ORGANIZATION_BLOCK "Cycle Execution"   // OB1, LAD
{ S7_Optimized_Access := 'FALSE' }
VERSION : 0.1
   VAR_TEMP
      TEMP0 : Byte;
      TEMP1 : Byte;
      TEMP2 : Byte;
      TEMP3 : Byte;
      TEMP4 : Byte;
      TEMP5 : Byte;
      TEMP6 : Int;
      TEMP7 : Int;
      TEMP8 : Int;
      TEMP9 : Date_And_Time;
      TEMP10 : DInt;
      TEMP11 : Int;
   END_VAR
   VAR_TEMP   // added for the SCL form of the ladder/FBD networks
      _w1 : Bool;
   END_VAR
BEGIN

REGION Network 1: -ALARMA
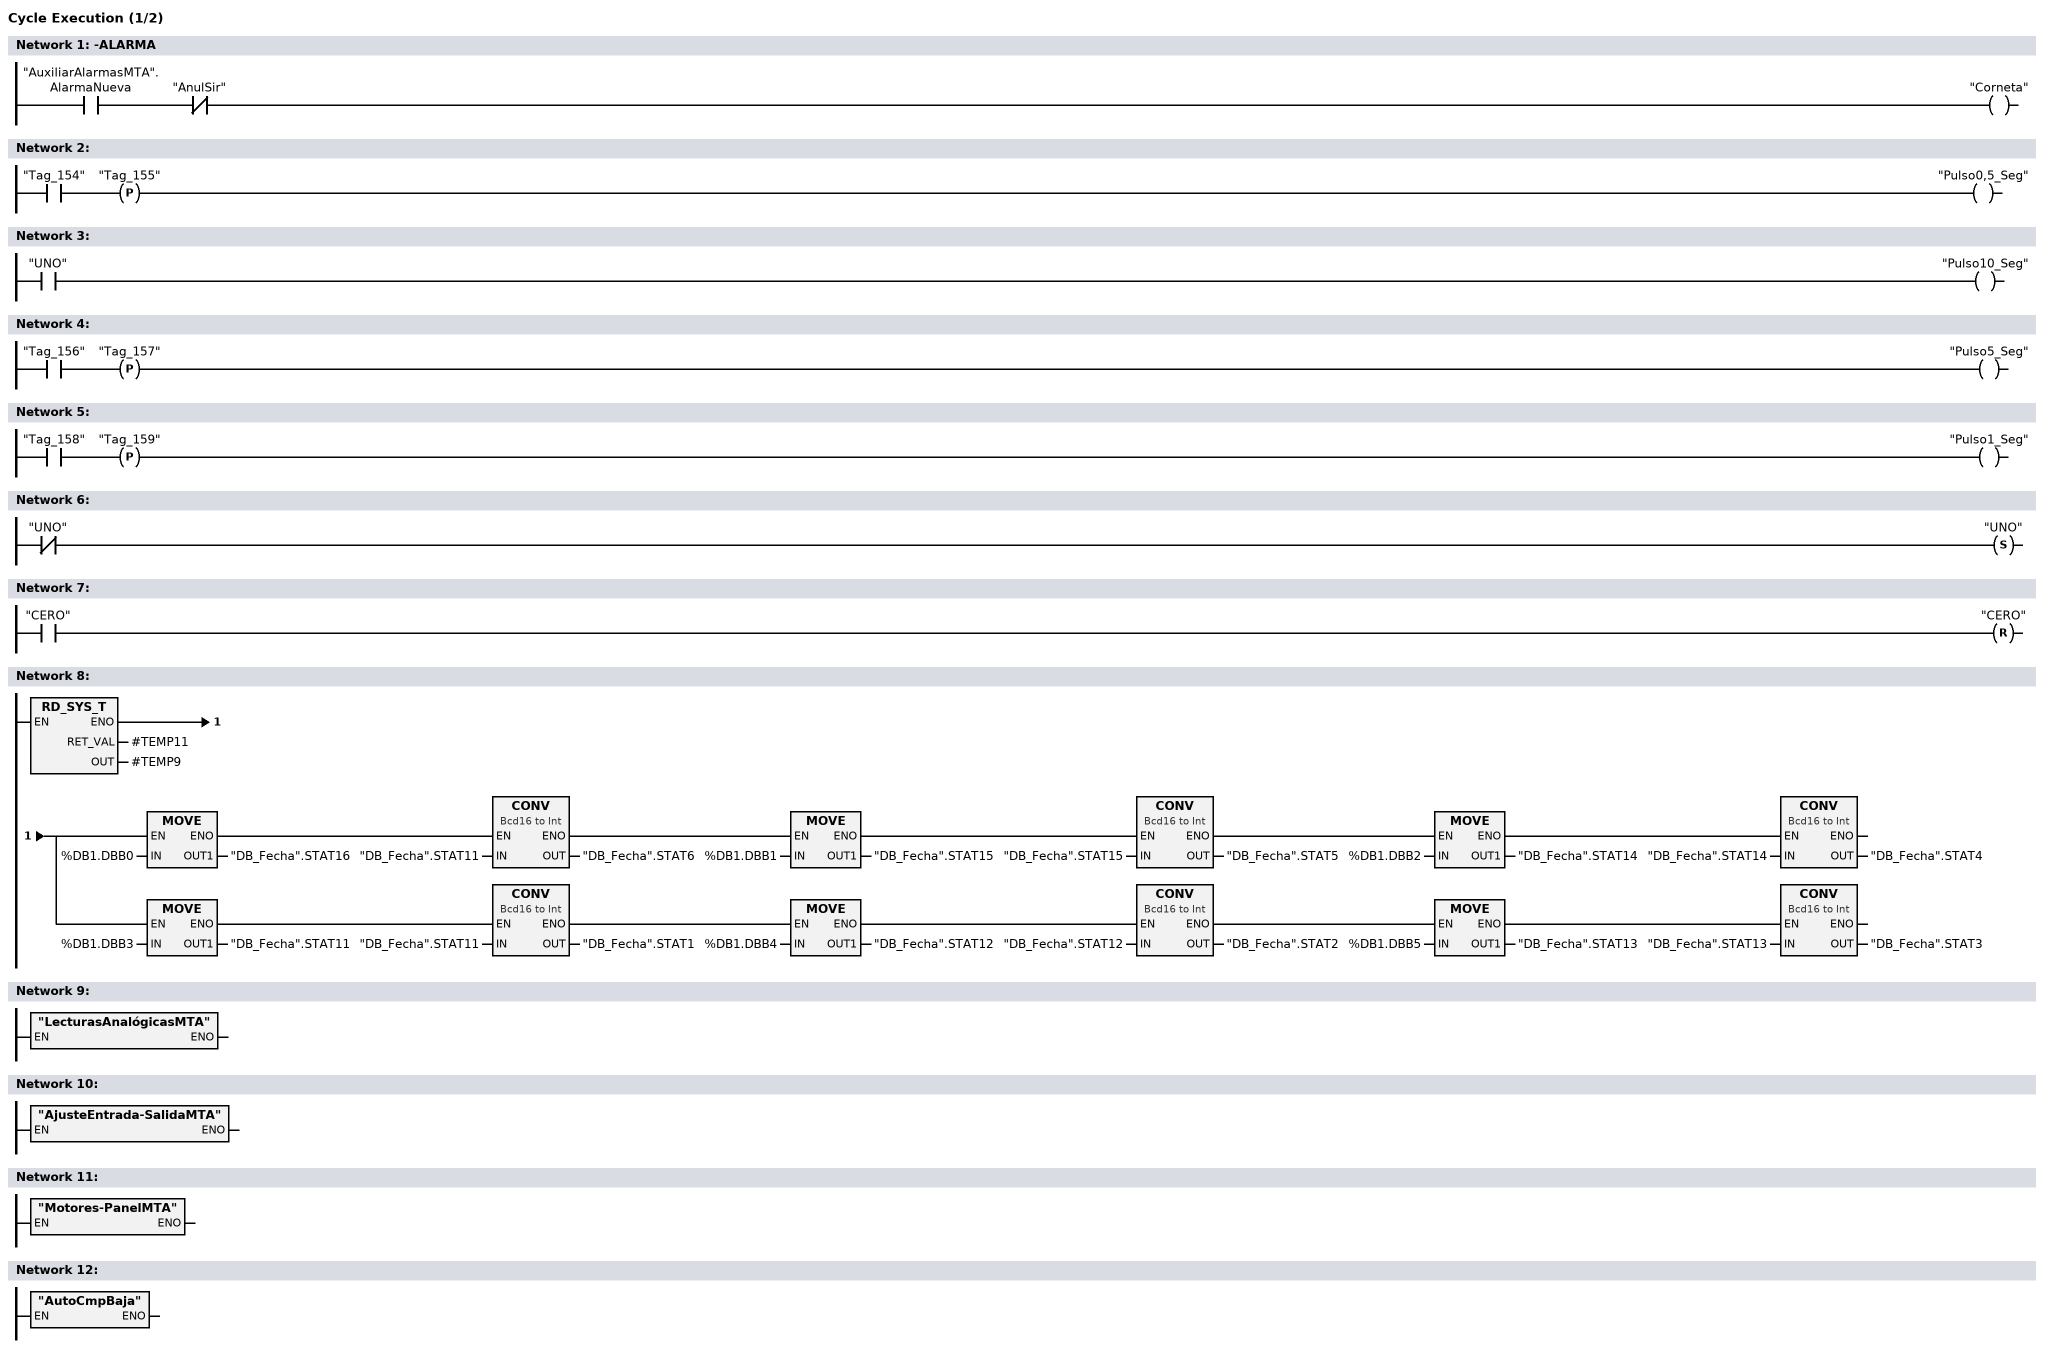
   RUNG wire#powerrail
      Contact( "AuxiliarAlarmasMTA".AlarmaNueva )
      I_Contact( "AnulSir" )
      Coil( "Corneta" )
   END_RUNG
   // the same network as SCL:
   "Corneta" := "AuxiliarAlarmasMTA".AlarmaNueva AND NOT "AnulSir";
END_REGION

REGION Network 2
   RUNG wire#powerrail
      Contact( "Tag_154" )
      P_Trig( "Tag_155" )
      Coil( "Pulso0,5_Seg" )
   END_RUNG
   // the same network as SCL:
   #_w1 := "Tag_154" AND NOT "Tag_155";   // rising edge
   "Tag_155" := "Tag_154";
   "Pulso0,5_Seg" := #_w1;
END_REGION

REGION Network 3
   RUNG wire#powerrail
      Contact( "UNO" )
      Coil( "Pulso10_Seg" )
   END_RUNG
   // the same network as SCL:
   "Pulso10_Seg" := "UNO";
END_REGION

REGION Network 4
   RUNG wire#powerrail
      Contact( "Tag_156" )
      P_Trig( "Tag_157" )
      Coil( "Pulso5_Seg" )
   END_RUNG
   // the same network as SCL:
   #_w1 := "Tag_156" AND NOT "Tag_157";   // rising edge
   "Tag_157" := "Tag_156";
   "Pulso5_Seg" := #_w1;
END_REGION

REGION Network 5
   RUNG wire#powerrail
      Contact( "Tag_158" )
      P_Trig( "Tag_159" )
      Coil( "Pulso1_Seg" )
   END_RUNG
   // the same network as SCL:
   #_w1 := "Tag_158" AND NOT "Tag_159";   // rising edge
   "Tag_159" := "Tag_158";
   "Pulso1_Seg" := #_w1;
END_REGION

REGION Network 6
   RUNG wire#powerrail
      I_Contact( "UNO" )
      S_Coil( "UNO" )
   END_RUNG
   // the same network as SCL:
   IF NOT "UNO" THEN "UNO" := TRUE; END_IF;
END_REGION

REGION Network 7
   RUNG wire#powerrail
      Contact( "CERO" )
      R_Coil( "CERO" )
   END_RUNG
   // the same network as SCL:
   IF "CERO" THEN "CERO" := FALSE; END_IF;
END_REGION

REGION Network 8
   // ENO of a box is taken as its EN; it also drops when the box reports an error
   #TEMP11 := RD_SYS_T(OUT => #TEMP9);
   "DB_Fecha".STAT16 := %DB1.DBB0;
   "DB_Fecha".STAT6 := BCD16_TO_INT("DB_Fecha".STAT11);
   "DB_Fecha".STAT15 := %DB1.DBB1;
   "DB_Fecha".STAT5 := BCD16_TO_INT("DB_Fecha".STAT15);
   "DB_Fecha".STAT14 := %DB1.DBB2;
   "DB_Fecha".STAT4 := BCD16_TO_INT("DB_Fecha".STAT14);
   "DB_Fecha".STAT11 := %DB1.DBB3;
   "DB_Fecha".STAT1 := BCD16_TO_INT("DB_Fecha".STAT11);
   "DB_Fecha".STAT12 := %DB1.DBB4;
   "DB_Fecha".STAT2 := BCD16_TO_INT("DB_Fecha".STAT12);
   "DB_Fecha".STAT13 := %DB1.DBB5;
   "DB_Fecha".STAT3 := BCD16_TO_INT("DB_Fecha".STAT13);
END_REGION

REGION Network 9
   RUNG wire#powerrail
      "LecturasAnalógicasMTA"()
   END_RUNG
   // the same network as SCL:
   "LecturasAnalógicasMTA"();
END_REGION

REGION Network 10
   RUNG wire#powerrail
      "AjusteEntrada-SalidaMTA"()
   END_RUNG
   // the same network as SCL:
   "AjusteEntrada-SalidaMTA"();
END_REGION

REGION Network 11
   RUNG wire#powerrail
      "Motores-PanelMTA"()
   END_RUNG
   // the same network as SCL:
   "Motores-PanelMTA"();
END_REGION

REGION Network 12
   RUNG wire#powerrail
      "AutoCmpBaja"()
   END_RUNG
   // the same network as SCL:
   "AutoCmpBaja"();
END_REGION

REGION Network 13
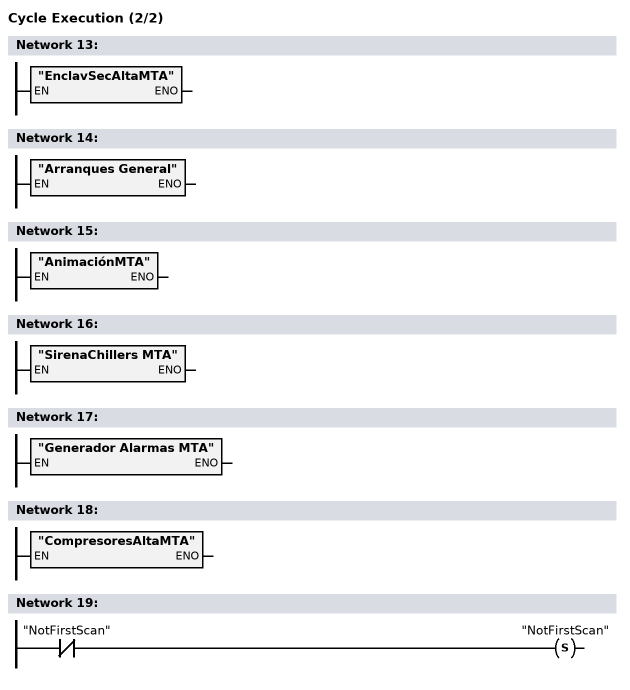
   RUNG wire#powerrail
      "EnclavSecAltaMTA"()
   END_RUNG
   // the same network as SCL:
   "EnclavSecAltaMTA"();
END_REGION

REGION Network 14
   RUNG wire#powerrail
      "Arranques General"()
   END_RUNG
   // the same network as SCL:
   "Arranques General"();
END_REGION

REGION Network 15
   RUNG wire#powerrail
      "AnimaciónMTA"()
   END_RUNG
   // the same network as SCL:
   "AnimaciónMTA"();
END_REGION

REGION Network 16
   RUNG wire#powerrail
      "SirenaChillers MTA"()
   END_RUNG
   // the same network as SCL:
   "SirenaChillers MTA"();
END_REGION

REGION Network 17
   RUNG wire#powerrail
      "Generador Alarmas MTA"()
   END_RUNG
   // the same network as SCL:
   "Generador Alarmas MTA"();
END_REGION

REGION Network 18
   RUNG wire#powerrail
      "CompresoresAltaMTA"()
   END_RUNG
   // the same network as SCL:
   "CompresoresAltaMTA"();
END_REGION

REGION Network 19
   RUNG wire#powerrail
      I_Contact( "NotFirstScan" )
      S_Coil( "NotFirstScan" )
   END_RUNG
   // the same network as SCL:
   IF NOT "NotFirstScan" THEN "NotFirstScan" := TRUE; END_IF;
END_REGION
END_ORGANIZATION_BLOCK

// folder: Alarmas

FUNCTION "SirenaChillers MTA" : Void   // FC7, LAD
{ S7_Optimized_Access := 'FALSE' }
VERSION : 0.1
BEGIN

REGION Network 1
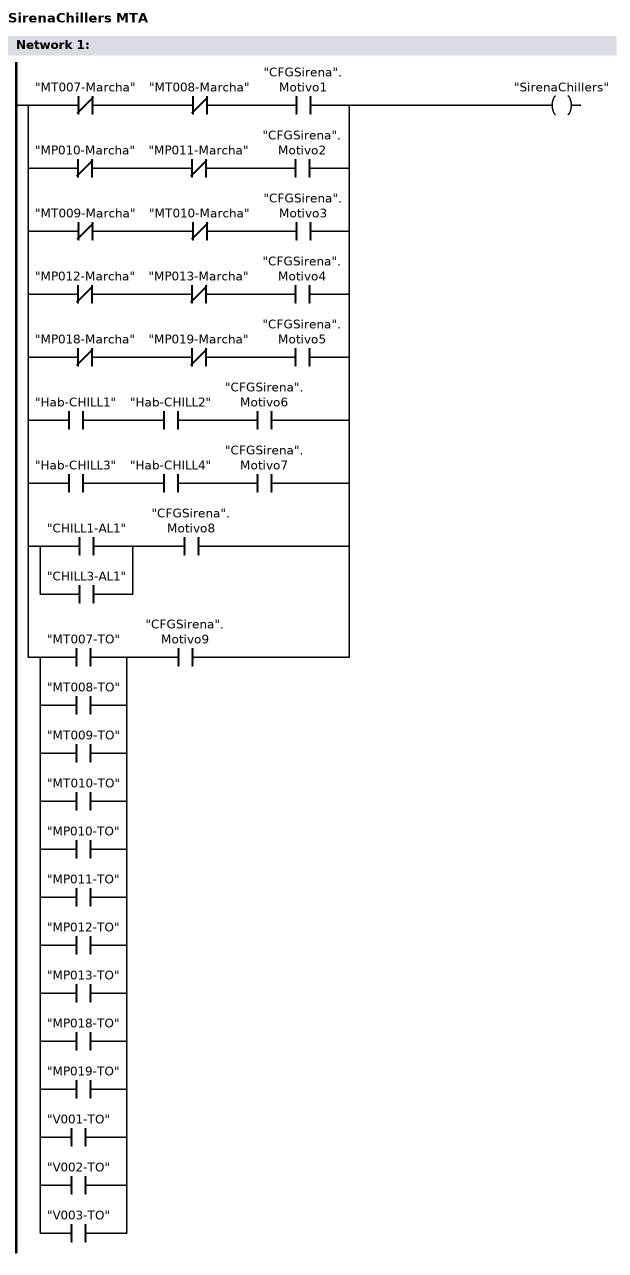
   RUNG wire#powerrail
      I_Contact( "MT007-Marcha" )
      I_Contact( "MT008-Marcha" )
      Contact( "CFGSirena".Motivo1 )
      wire#w1
      Coil( "SirenaChillers" )
   END_RUNG
   RUNG wire#powerrail
      I_Contact( "MP010-Marcha" )
      I_Contact( "MP011-Marcha" )
      Contact( "CFGSirena".Motivo2 )
   END_RUNG wire#w1
   RUNG wire#powerrail
      I_Contact( "MT009-Marcha" )
      I_Contact( "MT010-Marcha" )
      Contact( "CFGSirena".Motivo3 )
   END_RUNG wire#w1
   RUNG wire#powerrail
      I_Contact( "MP012-Marcha" )
      I_Contact( "MP013-Marcha" )
      Contact( "CFGSirena".Motivo4 )
   END_RUNG wire#w1
   RUNG wire#powerrail
      I_Contact( "MP018-Marcha" )
      I_Contact( "MP019-Marcha" )
      Contact( "CFGSirena".Motivo5 )
   END_RUNG wire#w1
   RUNG wire#powerrail
      Contact( "Hab-CHILL1" )
      Contact( "Hab-CHILL2" )
      Contact( "CFGSirena".Motivo6 )
   END_RUNG wire#w1
   RUNG wire#powerrail
      Contact( "Hab-CHILL3" )
      Contact( "Hab-CHILL4" )
      Contact( "CFGSirena".Motivo7 )
   END_RUNG wire#w1
   RUNG wire#powerrail
      Contact( "CHILL1-AL1" )
      wire#w2
      Contact( "CFGSirena".Motivo8 )
   END_RUNG wire#w1
   RUNG wire#powerrail
      Contact( "CHILL3-AL1" )
   END_RUNG wire#w2
   RUNG wire#powerrail
      Contact( "MT007-TO" )
      wire#w3
      Contact( "CFGSirena".Motivo9 )
   END_RUNG wire#w1
   RUNG wire#powerrail
      Contact( "MT008-TO" )
   END_RUNG wire#w3
   RUNG wire#powerrail
      Contact( "MT009-TO" )
   END_RUNG wire#w3
   RUNG wire#powerrail
      Contact( "MT010-TO" )
   END_RUNG wire#w3
   RUNG wire#powerrail
      Contact( "MP010-TO" )
   END_RUNG wire#w3
   RUNG wire#powerrail
      Contact( "MP011-TO" )
   END_RUNG wire#w3
   RUNG wire#powerrail
      Contact( "MP012-TO" )
   END_RUNG wire#w3
   RUNG wire#powerrail
      Contact( "MP013-TO" )
   END_RUNG wire#w3
   RUNG wire#powerrail
      Contact( "MP018-TO" )
   END_RUNG wire#w3
   RUNG wire#powerrail
      Contact( "MP019-TO" )
   END_RUNG wire#w3
   RUNG wire#powerrail
      Contact( "V001-TO" )
   END_RUNG wire#w3
   RUNG wire#powerrail
      Contact( "V002-TO" )
   END_RUNG wire#w3
   RUNG wire#powerrail
      Contact( "V003-TO" )
   END_RUNG wire#w3
   // the same network as SCL:
   "SirenaChillers" := (NOT "MT007-Marcha" AND NOT "MT008-Marcha" AND "CFGSirena".Motivo1) OR (NOT "MP010-Marcha" AND NOT "MP011-Marcha" AND "CFGSirena".Motivo2) OR (NOT "MT009-Marcha" AND NOT "MT010-Marcha" AND "CFGSirena".Motivo3) OR (NOT "MP012-Marcha" AND NOT "MP013-Marcha" AND "CFGSirena".Motivo4) OR (NOT "MP018-Marcha" AND NOT "MP019-Marcha" AND "CFGSirena".Motivo5) OR ("Hab-CHILL1" AND "Hab-CHILL2" AND "CFGSirena".Motivo6) OR ("Hab-CHILL3" AND "Hab-CHILL4" AND "CFGSirena".Motivo7) OR (("CHILL1-AL1" OR "CHILL3-AL1") AND "CFGSirena".Motivo8) OR (("MT007-TO" OR "MT008-TO" OR "MT009-TO" OR "MT010-TO" OR "MP010-TO" OR "MP011-TO" OR "MP012-TO" OR "MP013-TO" OR "MP018-TO" OR "MP019-TO" OR "V001-TO" OR "V002-TO" OR "V003-TO") AND "CFGSirena".Motivo9);
END_REGION
END_FUNCTION

FUNCTION "Generador Alarmas MTA" : Void   // FC8, LAD
{ S7_Optimized_Access := 'FALSE' }
VERSION : 0.1
   VAR_TEMP   // added for the SCL form of the ladder/FBD networks
      _w1 : Bool;
      _s5time1 : S5Time;
   END_VAR
BEGIN

REGION Network 1: Aviso 1 - Falla Conexión con sensor de Temperatura torres de Cavaleto
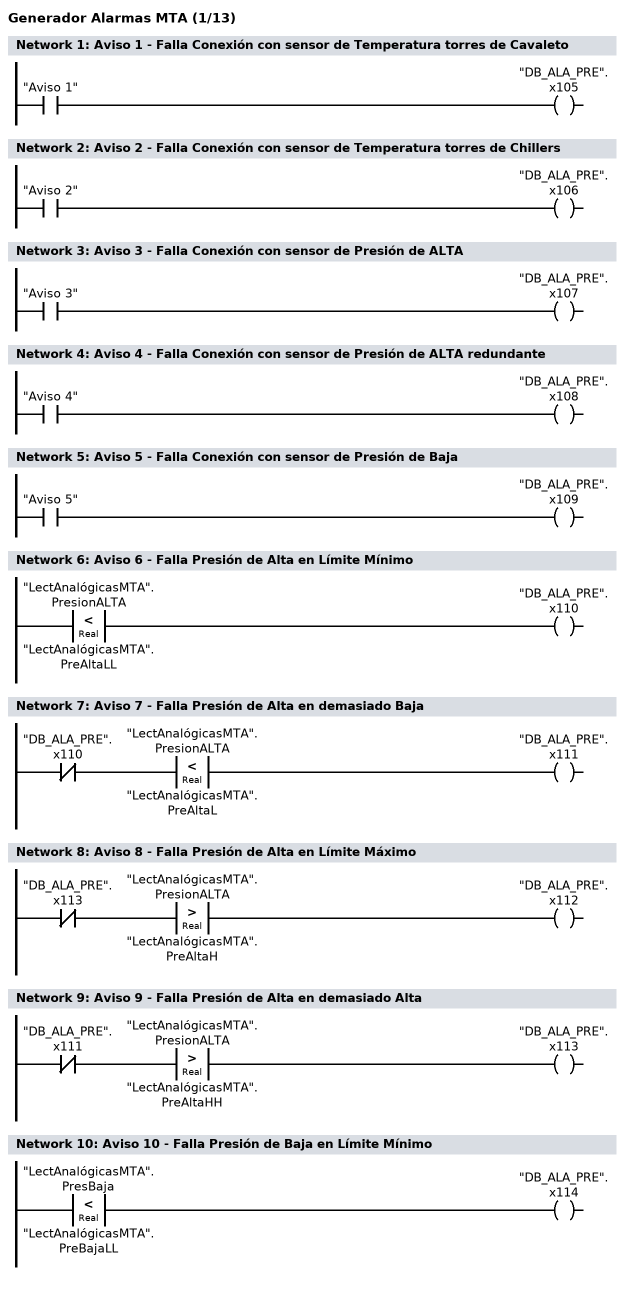
   RUNG wire#powerrail
      Contact( "Aviso 1" )
      Coil( "DB_ALA_PRE".x105 )
   END_RUNG
   // the same network as SCL:
   "DB_ALA_PRE".x105 := "Aviso 1";
END_REGION

REGION Network 2: Aviso 2 - Falla Conexión con sensor de Temperatura torres de Chillers
   RUNG wire#powerrail
      Contact( "Aviso 2" )
      Coil( "DB_ALA_PRE".x106 )
   END_RUNG
   // the same network as SCL:
   "DB_ALA_PRE".x106 := "Aviso 2";
END_REGION

REGION Network 3: Aviso 3 - Falla Conexión con sensor de Presión de ALTA
   RUNG wire#powerrail
      Contact( "Aviso 3" )
      Coil( "DB_ALA_PRE".x107 )
   END_RUNG
   // the same network as SCL:
   "DB_ALA_PRE".x107 := "Aviso 3";
END_REGION

REGION Network 4: Aviso 4 - Falla Conexión con sensor de Presión de ALTA redundante
   RUNG wire#powerrail
      Contact( "Aviso 4" )
      Coil( "DB_ALA_PRE".x108 )
   END_RUNG
   // the same network as SCL:
   "DB_ALA_PRE".x108 := "Aviso 4";
END_REGION

REGION Network 5: Aviso 5 - Falla Conexión con sensor de Presión de Baja
   RUNG wire#powerrail
      Contact( "Aviso 5" )
      Coil( "DB_ALA_PRE".x109 )
   END_RUNG
   // the same network as SCL:
   "DB_ALA_PRE".x109 := "Aviso 5";
END_REGION

REGION Network 6: Aviso 6 - Falla Presión de Alta en Límite Mínimo
   RUNG wire#powerrail
      { S7_Templates := "SrcType := Real" } LT_Contact(in1 := "LectAnalógicasMTA".PresionALTA, in2 := "LectAnalógicasMTA".PreAltaLL)
      Coil( "DB_ALA_PRE".x110 )
   END_RUNG
   // the same network as SCL:
   "DB_ALA_PRE".x110 := "LectAnalógicasMTA".PresionALTA < "LectAnalógicasMTA".PreAltaLL;
END_REGION

REGION Network 7: Aviso 7 - Falla Presión de Alta en demasiado Baja
   RUNG wire#powerrail
      I_Contact( "DB_ALA_PRE".x110 )
      { S7_Templates := "SrcType := Real" } LT_Contact(in1 := "LectAnalógicasMTA".PresionALTA, in2 := "LectAnalógicasMTA".PreAltaL)
      Coil( "DB_ALA_PRE".x111 )
   END_RUNG
   // the same network as SCL:
   "DB_ALA_PRE".x111 := NOT "DB_ALA_PRE".x110 AND ("LectAnalógicasMTA".PresionALTA < "LectAnalógicasMTA".PreAltaL);
END_REGION

REGION Network 8: Aviso 8 - Falla Presión de Alta en Límite Máximo
   RUNG wire#powerrail
      I_Contact( "DB_ALA_PRE".x113 )
      { S7_Templates := "SrcType := Real" } GT_Contact(in1 := "LectAnalógicasMTA".PresionALTA, in2 := "LectAnalógicasMTA".PreAltaH)
      Coil( "DB_ALA_PRE".x112 )
   END_RUNG
   // the same network as SCL:
   "DB_ALA_PRE".x112 := NOT "DB_ALA_PRE".x113 AND ("LectAnalógicasMTA".PresionALTA > "LectAnalógicasMTA".PreAltaH);
END_REGION

REGION Network 9: Aviso 9 - Falla Presión de Alta en demasiado Alta
   RUNG wire#powerrail
      I_Contact( "DB_ALA_PRE".x111 )
      { S7_Templates := "SrcType := Real" } GT_Contact(in1 := "LectAnalógicasMTA".PresionALTA, in2 := "LectAnalógicasMTA".PreAltaHH)
      Coil( "DB_ALA_PRE".x113 )
   END_RUNG
   // the same network as SCL:
   "DB_ALA_PRE".x113 := NOT "DB_ALA_PRE".x111 AND ("LectAnalógicasMTA".PresionALTA > "LectAnalógicasMTA".PreAltaHH);
END_REGION

REGION Network 10: Aviso 10 - Falla Presión de Baja en Límite Mínimo
   RUNG wire#powerrail
      { S7_Templates := "SrcType := Real" } LT_Contact(in1 := "LectAnalógicasMTA".PresBaja, in2 := "LectAnalógicasMTA".PreBajaLL)
      Coil( "DB_ALA_PRE".x114 )
   END_RUNG
   // the same network as SCL:
   "DB_ALA_PRE".x114 := "LectAnalógicasMTA".PresBaja < "LectAnalógicasMTA".PreBajaLL;
END_REGION

REGION Network 11: Aviso 11 - Falla Presión de Baja en demasiado Baja
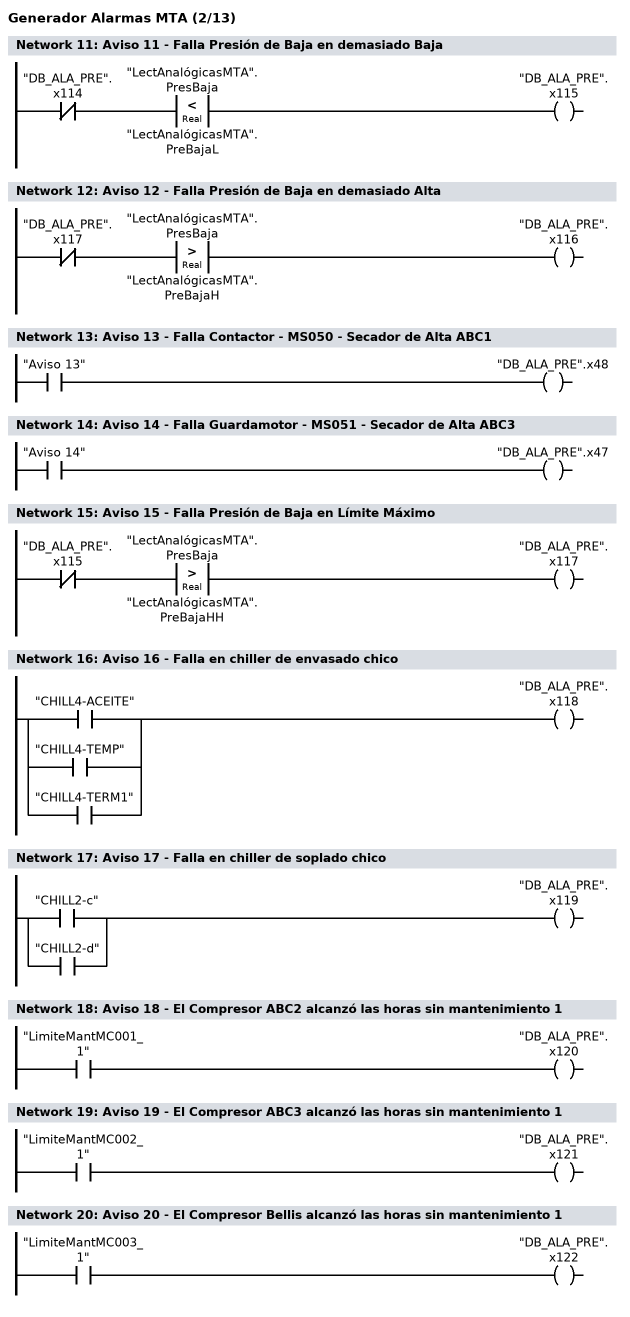
   RUNG wire#powerrail
      I_Contact( "DB_ALA_PRE".x114 )
      { S7_Templates := "SrcType := Real" } LT_Contact(in1 := "LectAnalógicasMTA".PresBaja, in2 := "LectAnalógicasMTA".PreBajaL)
      Coil( "DB_ALA_PRE".x115 )
   END_RUNG
   // the same network as SCL:
   "DB_ALA_PRE".x115 := NOT "DB_ALA_PRE".x114 AND ("LectAnalógicasMTA".PresBaja < "LectAnalógicasMTA".PreBajaL);
END_REGION

REGION Network 12: Aviso 12 - Falla Presión de Baja en demasiado Alta
   RUNG wire#powerrail
      I_Contact( "DB_ALA_PRE".x117 )
      { S7_Templates := "SrcType := Real" } GT_Contact(in1 := "LectAnalógicasMTA".PresBaja, in2 := "LectAnalógicasMTA".PreBajaH)
      Coil( "DB_ALA_PRE".x116 )
   END_RUNG
   // the same network as SCL:
   "DB_ALA_PRE".x116 := NOT "DB_ALA_PRE".x117 AND ("LectAnalógicasMTA".PresBaja > "LectAnalógicasMTA".PreBajaH);
END_REGION

REGION Network 13: Aviso 13 - Falla Contactor - MS050 - Secador de Alta ABC1
   RUNG wire#powerrail
      Contact( "Aviso 13" )
      Coil( "DB_ALA_PRE".x48 )
   END_RUNG
   // the same network as SCL:
   "DB_ALA_PRE".x48 := "Aviso 13";
END_REGION

REGION Network 14: Aviso 14 - Falla Guardamotor - MS051 - Secador de Alta ABC3
   RUNG wire#powerrail
      Contact( "Aviso 14" )
      Coil( "DB_ALA_PRE".x47 )
   END_RUNG
   // the same network as SCL:
   "DB_ALA_PRE".x47 := "Aviso 14";
END_REGION

REGION Network 15: Aviso 15 - Falla Presión de Baja en Límite Máximo
   RUNG wire#powerrail
      I_Contact( "DB_ALA_PRE".x115 )
      { S7_Templates := "SrcType := Real" } GT_Contact(in1 := "LectAnalógicasMTA".PresBaja, in2 := "LectAnalógicasMTA".PreBajaHH)
      Coil( "DB_ALA_PRE".x117 )
   END_RUNG
   // the same network as SCL:
   "DB_ALA_PRE".x117 := NOT "DB_ALA_PRE".x115 AND ("LectAnalógicasMTA".PresBaja > "LectAnalógicasMTA".PreBajaHH);
END_REGION

REGION Network 16: Aviso 16 - Falla en chiller de envasado chico
   RUNG wire#powerrail
      Contact( "CHILL4-ACEITE" )
      wire#w1
      Coil( "DB_ALA_PRE".x118 )
   END_RUNG
   RUNG wire#powerrail
      Contact( "CHILL4-TEMP" )
   END_RUNG wire#w1
   RUNG wire#powerrail
      Contact( "CHILL4-TERM1" )
   END_RUNG wire#w1
   // the same network as SCL:
   "DB_ALA_PRE".x118 := "CHILL4-ACEITE" OR "CHILL4-TEMP" OR "CHILL4-TERM1";
END_REGION

REGION Network 17: Aviso 17 - Falla en chiller de soplado chico
   RUNG wire#powerrail
      Contact( "CHILL2-c" )
      wire#w1
      Coil( "DB_ALA_PRE".x119 )
   END_RUNG
   RUNG wire#powerrail
      Contact( "CHILL2-d" )
   END_RUNG wire#w1
   // the same network as SCL:
   "DB_ALA_PRE".x119 := "CHILL2-c" OR "CHILL2-d";
END_REGION

REGION Network 18: Aviso 18 - El Compresor ABC2 alcanzó las horas sin mantenimiento 1
   RUNG wire#powerrail
      Contact( "LimiteMantMC001_1" )
      Coil( "DB_ALA_PRE".x120 )
   END_RUNG
   // the same network as SCL:
   "DB_ALA_PRE".x120 := "LimiteMantMC001_1";
END_REGION

REGION Network 19: Aviso 19 - El Compresor ABC3 alcanzó las horas sin mantenimiento 1
   RUNG wire#powerrail
      Contact( "LimiteMantMC002_1" )
      Coil( "DB_ALA_PRE".x121 )
   END_RUNG
   // the same network as SCL:
   "DB_ALA_PRE".x121 := "LimiteMantMC002_1";
END_REGION

REGION Network 20: Aviso 20 - El Compresor Bellis alcanzó las horas sin mantenimiento 1
   RUNG wire#powerrail
      Contact( "LimiteMantMC003_1" )
      Coil( "DB_ALA_PRE".x122 )
   END_RUNG
   // the same network as SCL:
   "DB_ALA_PRE".x122 := "LimiteMantMC003_1";
END_REGION

REGION Network 21: Aviso 21 - El Compresor ABC4 alcanzó las horas sin mantenimiento 1
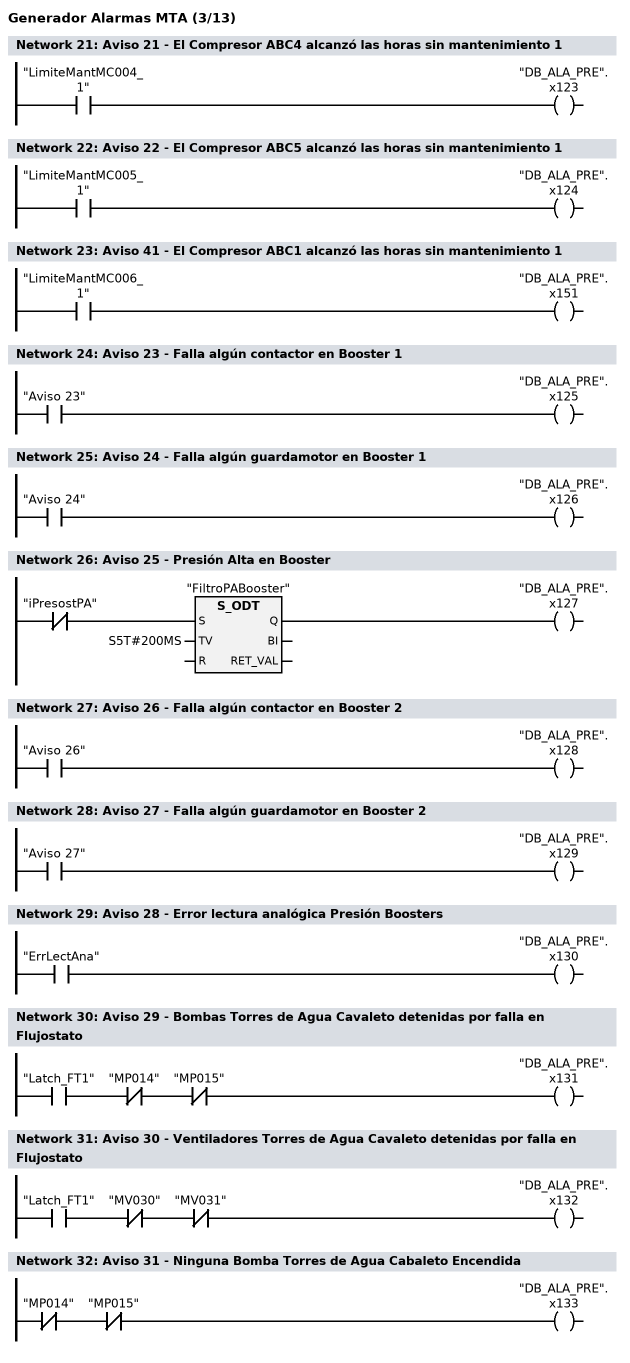
   RUNG wire#powerrail
      Contact( "LimiteMantMC004_1" )
      Coil( "DB_ALA_PRE".x123 )
   END_RUNG
   // the same network as SCL:
   "DB_ALA_PRE".x123 := "LimiteMantMC004_1";
END_REGION

REGION Network 22: Aviso 22 - El Compresor ABC5 alcanzó las horas sin mantenimiento 1
   RUNG wire#powerrail
      Contact( "LimiteMantMC005_1" )
      Coil( "DB_ALA_PRE".x124 )
   END_RUNG
   // the same network as SCL:
   "DB_ALA_PRE".x124 := "LimiteMantMC005_1";
END_REGION

REGION Network 23: Aviso 41 - El Compresor ABC1 alcanzó las horas sin mantenimiento 1
   RUNG wire#powerrail
      Contact( "LimiteMantMC006_1" )
      Coil( "DB_ALA_PRE".x151 )
   END_RUNG
   // the same network as SCL:
   "DB_ALA_PRE".x151 := "LimiteMantMC006_1";
END_REGION

REGION Network 24: Aviso 23 - Falla algún contactor en Booster 1
   RUNG wire#powerrail
      Contact( "Aviso 23" )
      Coil( "DB_ALA_PRE".x125 )
   END_RUNG
   // the same network as SCL:
   "DB_ALA_PRE".x125 := "Aviso 23";
END_REGION

REGION Network 25: Aviso 24 - Falla algún guardamotor en Booster 1
   RUNG wire#powerrail
      Contact( "Aviso 24" )
      Coil( "DB_ALA_PRE".x126 )
   END_RUNG
   // the same network as SCL:
   "DB_ALA_PRE".x126 := "Aviso 24";
END_REGION

REGION Network 26: Aviso 25 - Presión Alta en Booster
   RUNG wire#powerrail
      I_Contact( "iPresostPA" )
      S_ODT(T_NO := "FiltroPABooster", TV := S5T#200MS, R :=, BI =>, RET_VAL =>)
      Coil( "DB_ALA_PRE".x127 )
   END_RUNG
   // the same network as SCL:
   #_s5time1 := S_ODT(T_NO := "FiltroPABooster", S := NOT "iPresostPA", TV := S5T#200MS, Q => #_w1);
   "DB_ALA_PRE".x127 := #_w1;
END_REGION

REGION Network 27: Aviso 26 - Falla algún contactor en Booster 2
   RUNG wire#powerrail
      Contact( "Aviso 26" )
      Coil( "DB_ALA_PRE".x128 )
   END_RUNG
   // the same network as SCL:
   "DB_ALA_PRE".x128 := "Aviso 26";
END_REGION

REGION Network 28: Aviso 27 - Falla algún guardamotor en Booster 2
   RUNG wire#powerrail
      Contact( "Aviso 27" )
      Coil( "DB_ALA_PRE".x129 )
   END_RUNG
   // the same network as SCL:
   "DB_ALA_PRE".x129 := "Aviso 27";
END_REGION

REGION Network 29: Aviso 28 - Error lectura analógica Presión Boosters
   RUNG wire#powerrail
      Contact( "ErrLectAna" )
      Coil( "DB_ALA_PRE".x130 )
   END_RUNG
   // the same network as SCL:
   "DB_ALA_PRE".x130 := "ErrLectAna";
END_REGION

REGION Network 30: Aviso 29 - Bombas Torres de Agua Cavaleto detenidas por falla en Flujostato
   RUNG wire#powerrail
      Contact( "Latch_FT1" )
      I_Contact( "MP014" )
      I_Contact( "MP015" )
      Coil( "DB_ALA_PRE".x131 )
   END_RUNG
   // the same network as SCL:
   "DB_ALA_PRE".x131 := "Latch_FT1" AND NOT "MP014" AND NOT "MP015";
END_REGION

REGION Network 31: Aviso 30 - Ventiladores Torres de Agua Cavaleto detenidas por falla en Flujostato
   RUNG wire#powerrail
      Contact( "Latch_FT1" )
      I_Contact( "MV030" )
      I_Contact( "MV031" )
      Coil( "DB_ALA_PRE".x132 )
   END_RUNG
   // the same network as SCL:
   "DB_ALA_PRE".x132 := "Latch_FT1" AND NOT "MV030" AND NOT "MV031";
END_REGION

REGION Network 32: Aviso 31 - Ninguna Bomba Torres de Agua Cabaleto Encendida
   RUNG wire#powerrail
      I_Contact( "MP014" )
      I_Contact( "MP015" )
      Coil( "DB_ALA_PRE".x133 )
   END_RUNG
   // the same network as SCL:
   "DB_ALA_PRE".x133 := NOT "MP014" AND NOT "MP015";
END_REGION

REGION Network 33: Aviso 32 - Compresores Alta Detenidos por Flujostato Torres de Agua Cabaleto